(* Logix 5000 project; controller MV vendor 1 type 14 code 217 rev 31.11; software revision 31.00; part 33 of 53 *)
(* tags used below, declared in another part *)
   active : BOOL;
   Alarm_Reset : BOOL;
   CheckTimeMask : INT;
   CLOCK_system_set : BOOL;
   CLOCKsetvalues : DINT[7];
   colon_string : STRING;
   CurrentTime : DateTime;
   CWD : CHECKWORD_FLAGS;
   Default_Check_Time : DINT;
   FtoF_raw_input : REAL;
   FVHR26_3102 : PlantItem;   // Valve FVHR26_31/02
   FVHR26_3102_ALARM : ALARM_DIGITAL;
   FVHR26_3102_CL : ALIAS FOR RIO_Rack_2:14:I.Data.4;   // Valve FVHR26_31/02 Closed
   FVHR26_3102_DR : ALIAS FOR RIO_Rack_2:15:O.Data.18;   // Valve FVHR26_31/02 Drive
   FVHR26_3102_OP : ALIAS FOR RIO_Rack_2:14:I.Data.5;   // Valve FVHR26_31/02 Open
   FVHR26_3103 : PlantItem;   // Valve FVHR26_31/03
   FVHR26_3103_ALARM : ALARM_DIGITAL;
   FVHR26_3103_CL : ALIAS FOR RIO_Rack_2:14:I.Data.6;   // Valve FVHR26_31/03 Closed
   FVHR26_3103_DR : ALIAS FOR RIO_Rack_2:15:O.Data.19;   // Valve FVHR26_31/03 Drive
   FVHR26_3103_OP : ALIAS FOR RIO_Rack_2:14:I.Data.7;   // Valve FVHR26_31/03 Open
   FVHRCH201 : PlantItem;   // Valve FVHRCH201
   FVHRCH201_ALARM : ALARM_DIGITAL;
   FVHRCH201_CL : ALIAS FOR RIO_Rack_2:14:I.Data.10;   // Valve FVHRCH201 Closed
   FVHRCH201_DR : ALIAS FOR RIO_Rack_2:15:O.Data.21;   // Valve FVHRCH201 Drive
   FVHRCH201_OP : ALIAS FOR RIO_Rack_2:14:I.Data.11;   // Valve FVHRCH201 Open
   FVHRCH202 : PlantItem;   // Valve FVHRCH202
   FVHRCH202_ALARM : ALARM_DIGITAL;
   FVHRCH202_CL : ALIAS FOR RIO_Rack_2:14:I.Data.14;   // Valve FVHRCH202 Closed
   FVHRCH202_DR : ALIAS FOR RIO_Rack_2:15:O.Data.23;   // Valve FVHRCH202 Drive
   FVHRCH202_OP : ALIAS FOR RIO_Rack_2:14:I.Data.15;   // Valve FVHRCH202 Open
   FVHRCW01 : PlantItem;   // Valve FVHRCW01
   FVHRCW01_ALARM : ALARM_DIGITAL;
   FVHRCW01_CL : ALIAS FOR RIO_Rack_2:14:I.Data.12;   // Valve FVHRCW01 Closed
   FVHRCW01_DR : ALIAS FOR RIO_Rack_2:15:O.Data.22;   // Valve FVHRCW01 Drive
   FVHRCW01_OP : ALIAS FOR RIO_Rack_2:14:I.Data.13;   // Valve FVHRCW01 Open
   FVHRM01 : PlantItem;   // Valve FVHRM01
   FVHRM01_ALARM : ALARM_DIGITAL;
   FVHRM01_CL : ALIAS FOR RIO_Rack_2:13:I.Data.30;   // Valve FVHRM01 Closed
   FVHRM01_DR : ALIAS FOR RIO_Rack_2:15:O.Data.15;   // Valve FVHRM01 Drive
   FVHRM01_OP : ALIAS FOR RIO_Rack_2:13:I.Data.31;   // Valve FVHRM01 Open
   FVHRM02 : PlantItem;   // Valve FVHRM02
   FVHRM02_ALARM : ALARM_DIGITAL;
   FVHRM02_CL : ALIAS FOR RIO_Rack_2:14:I.Data.0;   // Valve FVHRM02 Closed
   FVHRM02_DR : ALIAS FOR RIO_Rack_2:15:O.Data.16;   // Valve FVHRM02 Drive
   FVHRM02_OP : ALIAS FOR RIO_Rack_2:14:I.Data.1;   // Valve FVHRM02 Open
   FVHRM03 : PlantItem;   // Valve FVHRM03
   FVHRM03_ALARM : ALARM_DIGITAL;
   FVHRM03_CL : ALIAS FOR RIO_Rack_2:14:I.Data.8;   // Valve FVHRM03 Closed
   FVHRM03_DR : ALIAS FOR RIO_Rack_2:15:O.Data.20;   // Valve FVHRM03 Drive
   FVHRM03_OP : ALIAS FOR RIO_Rack_2:14:I.Data.9;   // Valve FVHRM03 Open
   FVHRM04 : PlantItem;   // Valve FVHRM04
   FVHRM04_ALARM : ALARM_DIGITAL;
   FVHRM04_CL : ALIAS FOR RIO_Rack_2:13:I.Data.12;   // Valve FVHRM04 Closed
   FVHRM04_DR : ALIAS FOR RIO_Rack_2:15:O.Data.6;   // Valve FVHRM04 Drive
   FVHRM04_OP : ALIAS FOR RIO_Rack_2:13:I.Data.13;   // Valve FVHRM04 Open
   FVHRMD01 : PlantItem;   // Valve FVHRMD01
   FVHRMD01_ALARM : ALARM_DIGITAL;
   FVHRMD01_CL : ALIAS FOR RIO_Rack_2:13:I.Data.14;   // Valve FVHRMD01 Closed
   FVHRMD01_DR : ALIAS FOR RIO_Rack_2:15:O.Data.7;   // Valve FVHRMD01 Drive
   FVHRMD01_OP : ALIAS FOR RIO_Rack_2:13:I.Data.15;   // Valve FVHRMD01 Open
   hr_string : STRING;
   IGI_TestBit : BOOL;
   Item_Faults_Are_Latched : BOOL;
   Item_Simulation_Flag : BOOL;
   ItoF_raw_input : INT;
   mn_string : STRING;
   MV_DayOfWeek : DINT;
   MV_DayOfWeekONS : BOOL;
   MV_SFile : INT[255];   // SLC Equivalent System File, So Original Code Can Remain
   One_Second_One_Scan : ALIAS FOR One_Second_1_scan;
   result_string : STRING;
   scale_analog_int : DINT;
   scale_analog_result : REAL;
   scale_eu_max : REAL;
   scale_eu_min : REAL;
   scale_raw_input : REAL;
   scale_raw_max : REAL;
   scale_raw_min : REAL;
   scale_routine_active : BOOL;
   scale_temp : REAL;
   se_string : STRING;
   seconds_input_DINT : DINT;
   temp : INT;
   temp_hr : INT;
   temp_mn : INT;
   temp_se : INT;
   zero_string : STRING;
(* MC_Common, continued *)

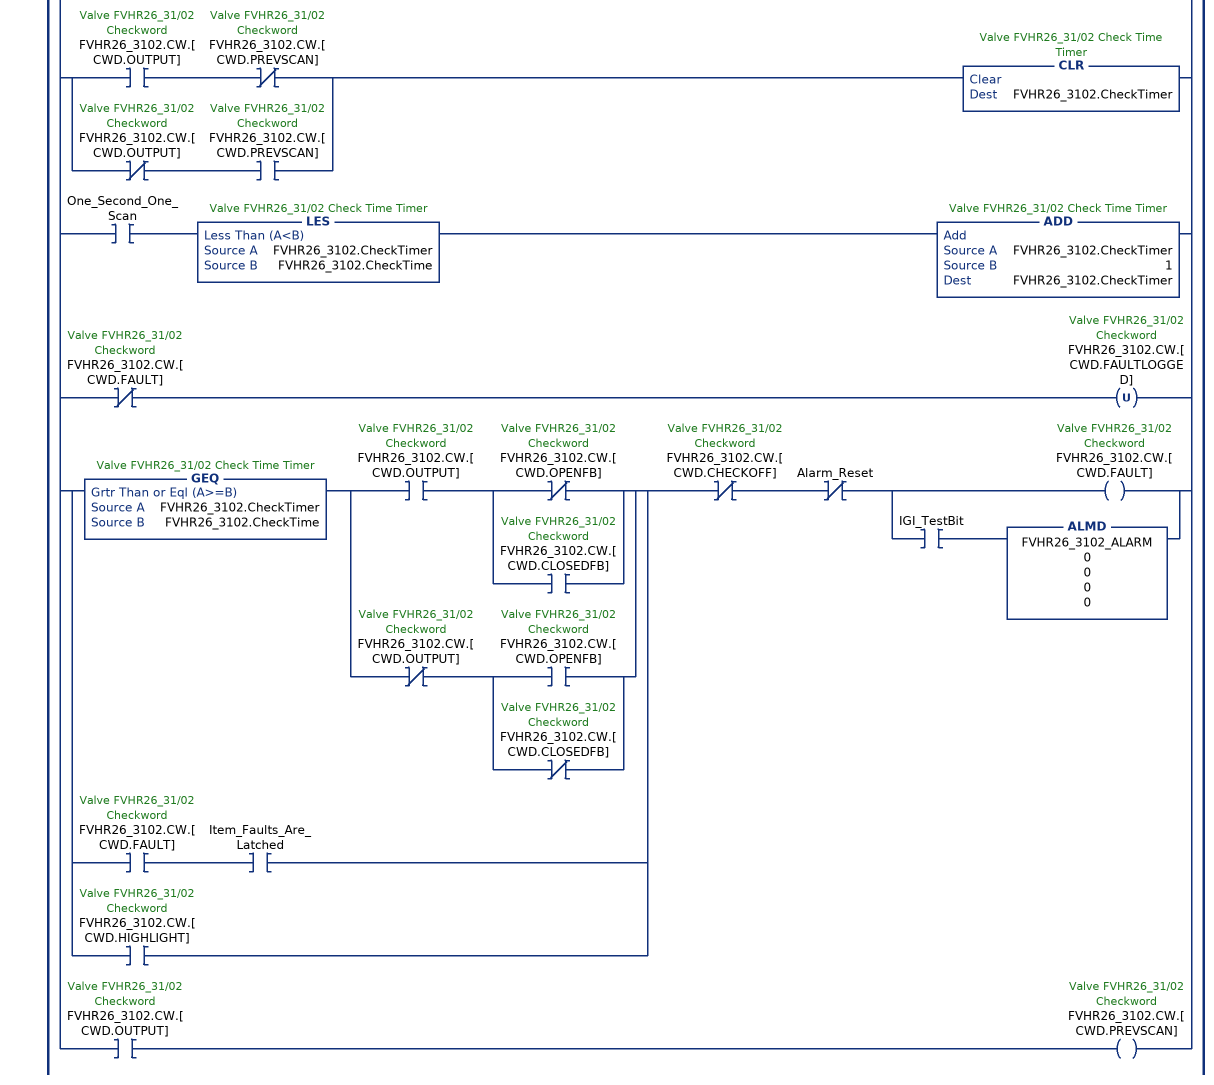
   [picture p757: MC_Common/MC_Valves rungs 79-79]
   79: [NEQ(FVHR26_3102.DriveBits,0) OTE(FVHR26_3102.CW.[CWD.AUTODRV]) ,[XIC(FVHR26_3102.CW.[CWD.AUTODRV]) XIO(FVHR26_3102.CW.[CWD.MANUAL]) ,XIC(FVHR26_3102.CW.[CWD.MANDRV]) XIC(FVHR26_3102.CW.[CWD.MANUAL]) ] OTE(FVHR26_3102.CW.[CWD.OUTPUT]) ,XIC(FVHR26_3102.CW.[CWD.OUTPUT]) OTE(FVHR26_3102_DR) ,XIC(S:FS) [OTU(FVHR26_3102.CW.[CWD.MANUAL]) ,LEQ(FVHR26_3102.CheckTime,0) MOV(Default_Check_Time,FVHR26_3102.CheckTime) ] ,[[XIC(FVHR26_3102_OP) XIO(Item_Simulation_Flag) ,XIC(Item_Simulation_Flag) XIC(FVHR26_3102.CW.[CWD.OUTPUT]) XIO(FVHR26_3102.CW.[CWD.SIMFAIL]) ] OTE(FVHR26_3102.CW.[CWD.OPENFB]) ,[XIC(FVHR26_3102_CL) XIO(Item_Simulation_Flag) ,XIC(Item_Simulation_Flag) XIO(FVHR26_3102.CW.[CWD.OUTPUT]) XIO(FVHR26_3102.CW.[CWD.SIMFAIL]) ] OTE(FVHR26_3102.CW.[CWD.CLOSEDFB]) ] ,[XIC(FVHR26_3102.CW.[CWD.OUTPUT]) XIO(FVHR26_3102.CW.[CWD.PREVSCAN]) ,XIO(FVHR26_3102.CW.[CWD.OUTPUT]) XIC(FVHR26_3102.CW.[CWD.PREVSCAN]) ] CLR(FVHR26_3102.CheckTimer) ,XIC(One_Second_One_Scan) LES(FVHR26_3102.CheckTimer,FVHR26_3102.CheckTime) ADD(FVHR26_3102.CheckTimer,1,FVHR26_3102.CheckTimer) ,XIO(FVHR26_3102.CW.[CWD.FAULT]) OTU(FVHR26_3102.CW.[CWD.FAULTLOGGED]) ,[GEQ(FVHR26_3102.CheckTimer,FVHR26_3102.CheckTime) [XIC(FVHR26_3102.CW.[CWD.OUTPUT]) [XIO(FVHR26_3102.CW.[CWD.OPENFB]) ,XIC(FVHR26_3102.CW.[CWD.CLOSEDFB]) ] ,XIO(FVHR26_3102.CW.[CWD.OUTPUT]) [XIC(FVHR26_3102.CW.[CWD.OPENFB]) ,XIO(FVHR26_3102.CW.[CWD.CLOSEDFB]) ] ] ,XIC(FVHR26_3102.CW.[CWD.FAULT]) XIC(Item_Faults_Are_Latched) ,XIC(FVHR26_3102.CW.[CWD.HIGHLIGHT]) ] XIO(FVHR26_3102.CW.[CWD.CHECKOFF]) XIO(Alarm_Reset) [OTE(FVHR26_3102.CW.[CWD.FAULT]) ,XIC(IGI_TestBit) ALMD(FVHR26_3102_ALARM,0,0,0,0) ] ,XIC(FVHR26_3102.CW.[CWD.OUTPUT]) OTE(FVHR26_3102.CW.[CWD.PREVSCAN]) ];
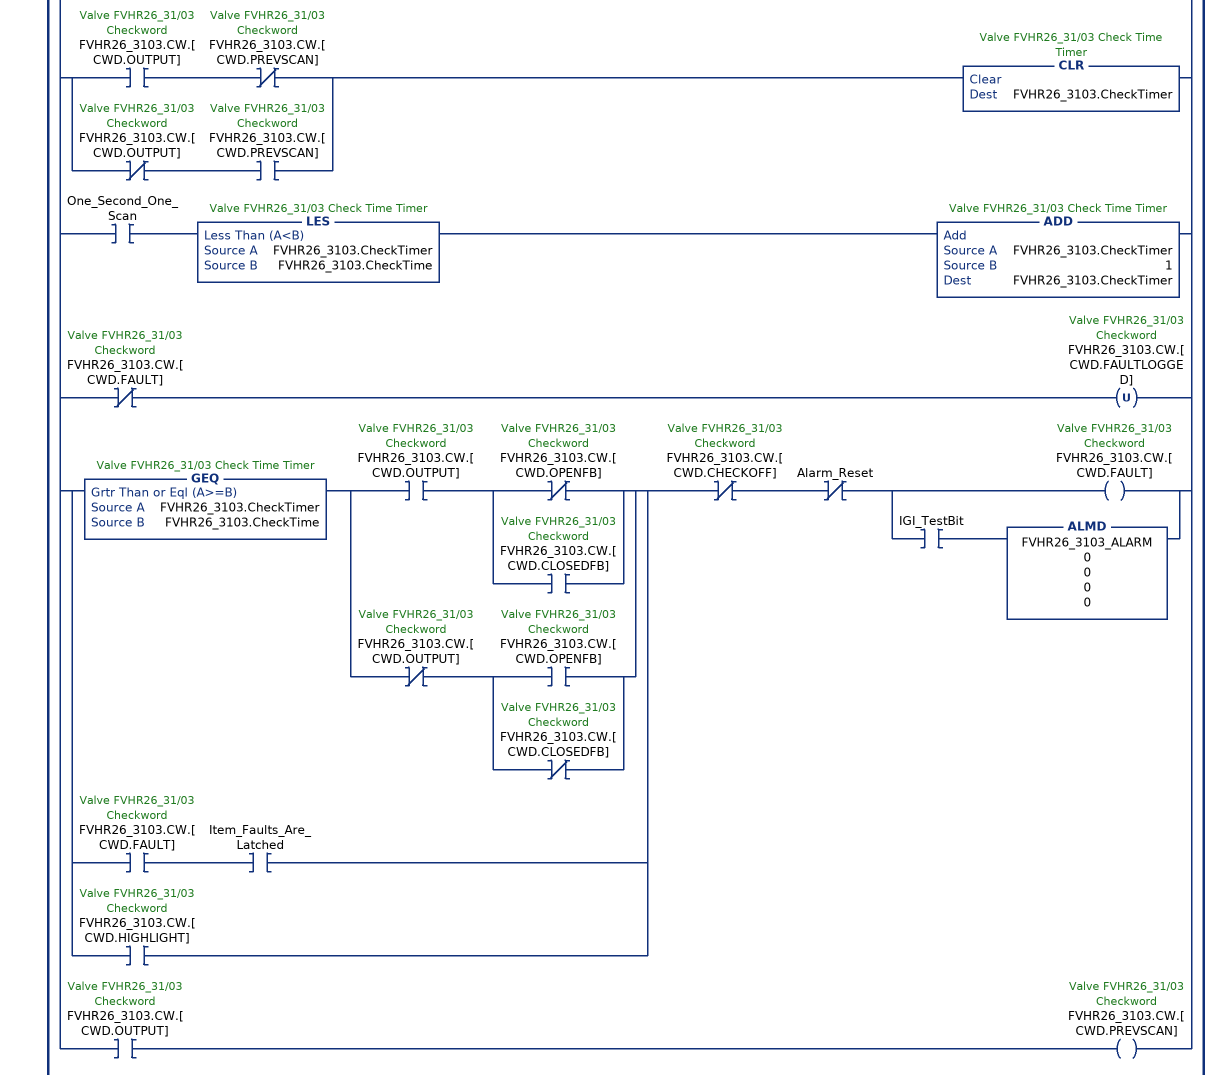
   80: [NEQ(FVHR26_3103.DriveBits,0) OTE(FVHR26_3103.CW.[CWD.AUTODRV]) ,[XIC(FVHR26_3103.CW.[CWD.AUTODRV]) XIO(FVHR26_3103.CW.[CWD.MANUAL]) ,XIC(FVHR26_3103.CW.[CWD.MANDRV]) XIC(FVHR26_3103.CW.[CWD.MANUAL]) ] OTE(FVHR26_3103.CW.[CWD.OUTPUT]) ,XIC(FVHR26_3103.CW.[CWD.OUTPUT]) OTE(FVHR26_3103_DR) ,XIC(S:FS) [OTU(FVHR26_3103.CW.[CWD.MANUAL]) ,LEQ(FVHR26_3103.CheckTime,0) MOV(Default_Check_Time,FVHR26_3103.CheckTime) ] ,[[XIC(FVHR26_3103_OP) XIO(Item_Simulation_Flag) ,XIC(Item_Simulation_Flag) XIC(FVHR26_3103.CW.[CWD.OUTPUT]) XIO(FVHR26_3103.CW.[CWD.SIMFAIL]) ] OTE(FVHR26_3103.CW.[CWD.OPENFB]) ,[XIC(FVHR26_3103_CL) XIO(Item_Simulation_Flag) ,XIC(Item_Simulation_Flag) XIO(FVHR26_3103.CW.[CWD.OUTPUT]) XIO(FVHR26_3103.CW.[CWD.SIMFAIL]) ] OTE(FVHR26_3103.CW.[CWD.CLOSEDFB]) ] ,[XIC(FVHR26_3103.CW.[CWD.OUTPUT]) XIO(FVHR26_3103.CW.[CWD.PREVSCAN]) ,XIO(FVHR26_3103.CW.[CWD.OUTPUT]) XIC(FVHR26_3103.CW.[CWD.PREVSCAN]) ] CLR(FVHR26_3103.CheckTimer) ,XIC(One_Second_One_Scan) LES(FVHR26_3103.CheckTimer,FVHR26_3103.CheckTime) ADD(FVHR26_3103.CheckTimer,1,FVHR26_3103.CheckTimer) ,XIO(FVHR26_3103.CW.[CWD.FAULT]) OTU(FVHR26_3103.CW.[CWD.FAULTLOGGED]) ,[GEQ(FVHR26_3103.CheckTimer,FVHR26_3103.CheckTime) [XIC(FVHR26_3103.CW.[CWD.OUTPUT]) [XIO(FVHR26_3103.CW.[CWD.OPENFB]) ,XIC(FVHR26_3103.CW.[CWD.CLOSEDFB]) ] ,XIO(FVHR26_3103.CW.[CWD.OUTPUT]) [XIC(FVHR26_3103.CW.[CWD.OPENFB]) ,XIO(FVHR26_3103.CW.[CWD.CLOSEDFB]) ] ] ,XIC(FVHR26_3103.CW.[CWD.FAULT]) XIC(Item_Faults_Are_Latched) ,XIC(FVHR26_3103.CW.[CWD.HIGHLIGHT]) ] XIO(FVHR26_3103.CW.[CWD.CHECKOFF]) XIO(Alarm_Reset) [OTE(FVHR26_3103.CW.[CWD.FAULT]) ,XIC(IGI_TestBit) ALMD(FVHR26_3103_ALARM,0,0,0,0) ] ,XIC(FVHR26_3103.CW.[CWD.OUTPUT]) OTE(FVHR26_3103.CW.[CWD.PREVSCAN]) ];
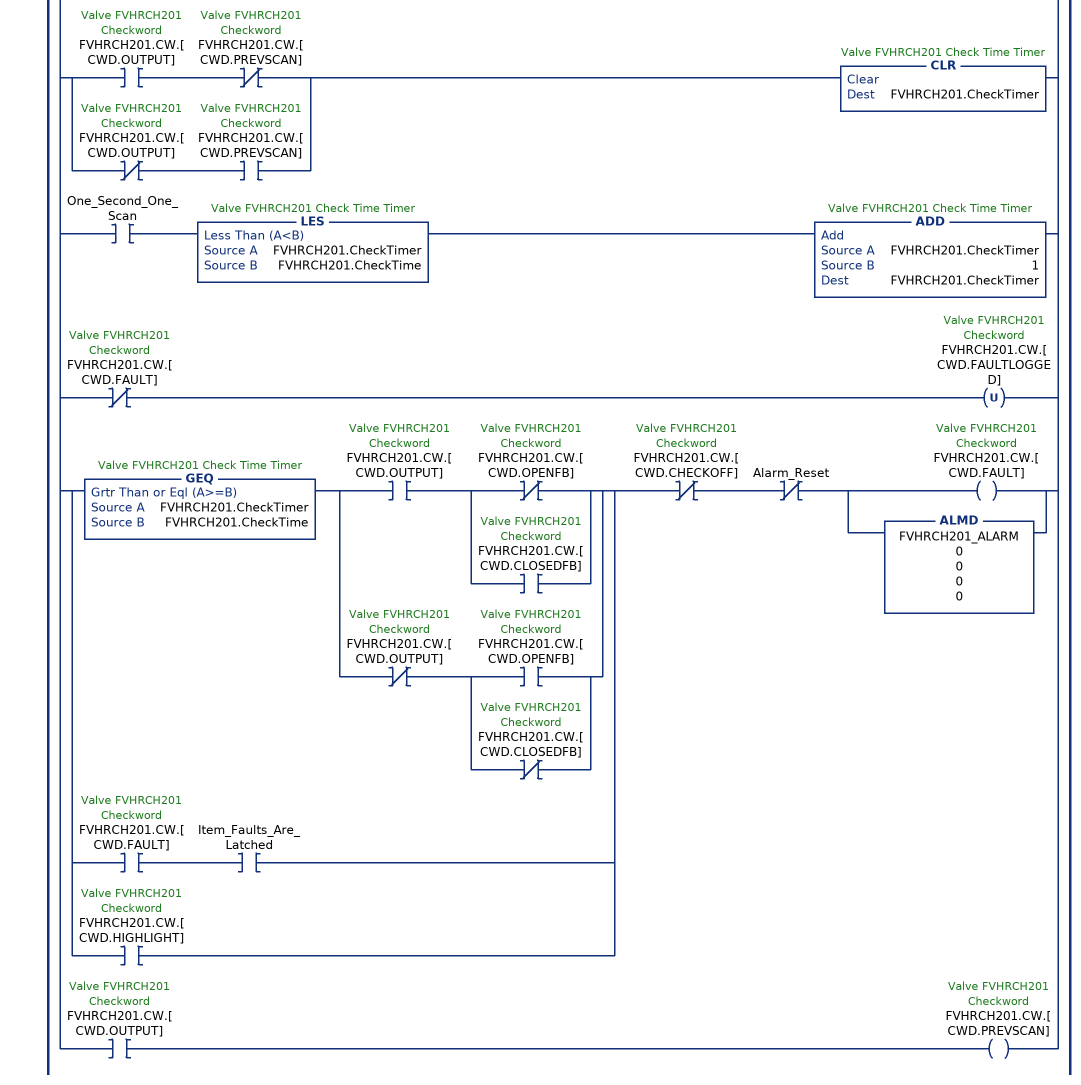
   81: [NEQ(FVHRCH201.DriveBits,0) OTE(FVHRCH201.CW.[CWD.AUTODRV]) ,[XIC(FVHRCH201.CW.[CWD.AUTODRV]) XIO(FVHRCH201.CW.[CWD.MANUAL]) ,XIC(FVHRCH201.CW.[CWD.MANDRV]) XIC(FVHRCH201.CW.[CWD.MANUAL]) ] OTE(FVHRCH201.CW.[CWD.OUTPUT]) ,XIC(FVHRCH201.CW.[CWD.OUTPUT]) OTE(FVHRCH201_DR) ,XIC(S:FS) [OTU(FVHRCH201.CW.[CWD.MANUAL]) ,LEQ(FVHRCH201.CheckTime,0) MOV(Default_Check_Time,FVHRCH201.CheckTime) ] ,[[XIC(FVHRCH201_OP) XIO(Item_Simulation_Flag) ,XIC(Item_Simulation_Flag) XIC(FVHRCH201.CW.[CWD.OUTPUT]) XIO(FVHRCH201.CW.[CWD.SIMFAIL]) ] OTE(FVHRCH201.CW.[CWD.OPENFB]) ,[XIC(FVHRCH201_CL) XIO(Item_Simulation_Flag) ,XIC(Item_Simulation_Flag) XIO(FVHRCH201.CW.[CWD.OUTPUT]) XIO(FVHRCH201.CW.[CWD.SIMFAIL]) ] OTE(FVHRCH201.CW.[CWD.CLOSEDFB]) ] ,[XIC(FVHRCH201.CW.[CWD.OUTPUT]) XIO(FVHRCH201.CW.[CWD.PREVSCAN]) ,XIO(FVHRCH201.CW.[CWD.OUTPUT]) XIC(FVHRCH201.CW.[CWD.PREVSCAN]) ] CLR(FVHRCH201.CheckTimer) ,XIC(One_Second_One_Scan) LES(FVHRCH201.CheckTimer,FVHRCH201.CheckTime) ADD(FVHRCH201.CheckTimer,1,FVHRCH201.CheckTimer) ,XIO(FVHRCH201.CW.[CWD.FAULT]) OTU(FVHRCH201.CW.[CWD.FAULTLOGGED]) ,[GEQ(FVHRCH201.CheckTimer,FVHRCH201.CheckTime) [XIC(FVHRCH201.CW.[CWD.OUTPUT]) [XIO(FVHRCH201.CW.[CWD.OPENFB]) ,XIC(FVHRCH201.CW.[CWD.CLOSEDFB]) ] ,XIO(FVHRCH201.CW.[CWD.OUTPUT]) [XIC(FVHRCH201.CW.[CWD.OPENFB]) ,XIO(FVHRCH201.CW.[CWD.CLOSEDFB]) ] ] ,XIC(FVHRCH201.CW.[CWD.FAULT]) XIC(Item_Faults_Are_Latched) ,XIC(FVHRCH201.CW.[CWD.HIGHLIGHT]) ] XIO(FVHRCH201.CW.[CWD.CHECKOFF]) XIO(Alarm_Reset) [OTE(FVHRCH201.CW.[CWD.FAULT]) ,ALMD(FVHRCH201_ALARM,0,0,0,0) ] ,XIC(FVHRCH201.CW.[CWD.OUTPUT]) OTE(FVHRCH201.CW.[CWD.PREVSCAN]) ];
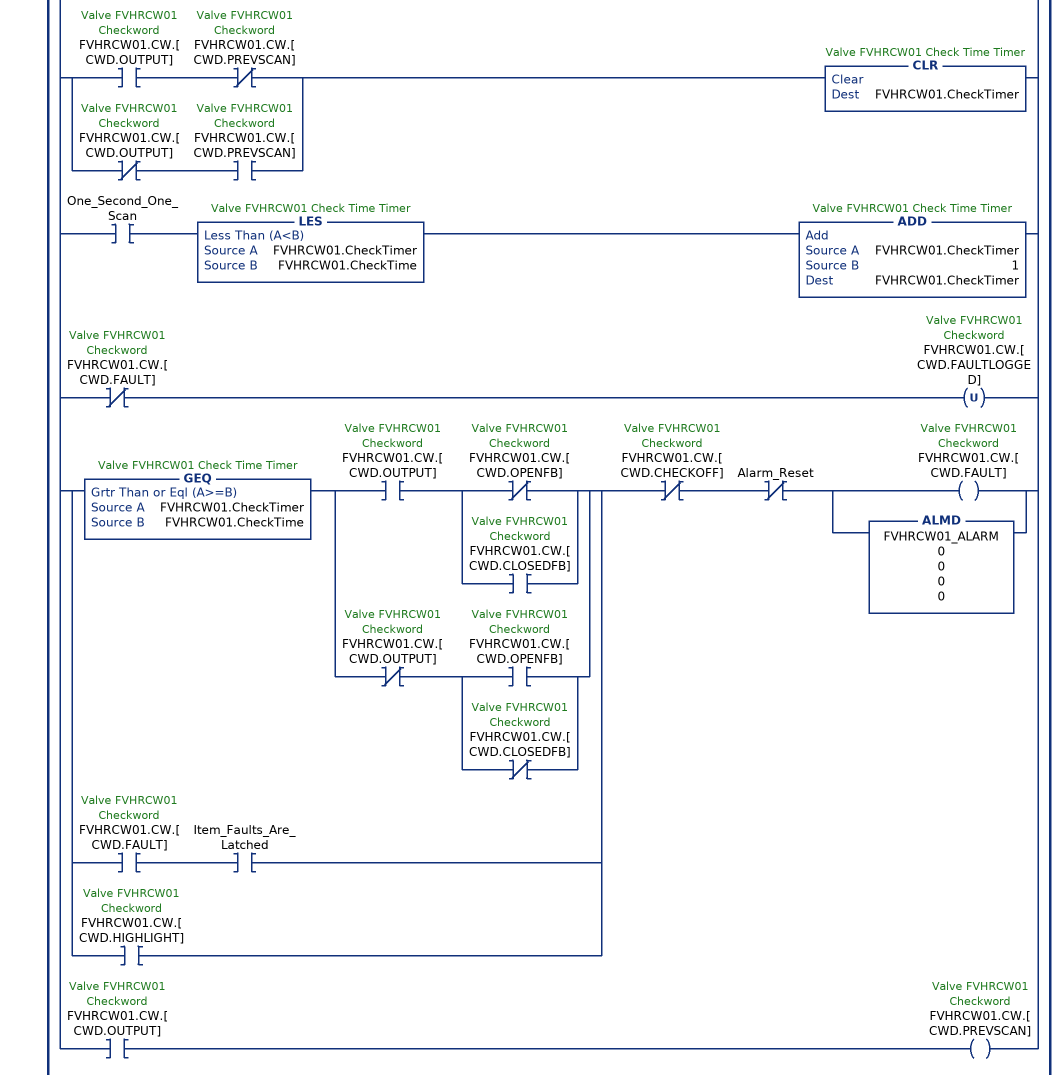
   82: [NEQ(FVHRCW01.DriveBits,0) OTE(FVHRCW01.CW.[CWD.AUTODRV]) ,[XIC(FVHRCW01.CW.[CWD.AUTODRV]) XIO(FVHRCW01.CW.[CWD.MANUAL]) ,XIC(FVHRCW01.CW.[CWD.MANDRV]) XIC(FVHRCW01.CW.[CWD.MANUAL]) ] OTE(FVHRCW01.CW.[CWD.OUTPUT]) ,XIC(FVHRCW01.CW.[CWD.OUTPUT]) OTE(FVHRCW01_DR) ,XIC(S:FS) [OTU(FVHRCW01.CW.[CWD.MANUAL]) ,LEQ(FVHRCW01.CheckTime,0) MOV(Default_Check_Time,FVHRCW01.CheckTime) ] ,[[XIC(FVHRCW01_OP) XIO(Item_Simulation_Flag) ,XIC(Item_Simulation_Flag) XIC(FVHRCW01.CW.[CWD.OUTPUT]) XIO(FVHRCW01.CW.[CWD.SIMFAIL]) ] OTE(FVHRCW01.CW.[CWD.OPENFB]) ,[XIC(FVHRCW01_CL) XIO(Item_Simulation_Flag) ,XIC(Item_Simulation_Flag) XIO(FVHRCW01.CW.[CWD.OUTPUT]) XIO(FVHRCW01.CW.[CWD.SIMFAIL]) ] OTE(FVHRCW01.CW.[CWD.CLOSEDFB]) ] ,[XIC(FVHRCW01.CW.[CWD.OUTPUT]) XIO(FVHRCW01.CW.[CWD.PREVSCAN]) ,XIO(FVHRCW01.CW.[CWD.OUTPUT]) XIC(FVHRCW01.CW.[CWD.PREVSCAN]) ] CLR(FVHRCW01.CheckTimer) ,XIC(One_Second_One_Scan) LES(FVHRCW01.CheckTimer,FVHRCW01.CheckTime) ADD(FVHRCW01.CheckTimer,1,FVHRCW01.CheckTimer) ,XIO(FVHRCW01.CW.[CWD.FAULT]) OTU(FVHRCW01.CW.[CWD.FAULTLOGGED]) ,[GEQ(FVHRCW01.CheckTimer,FVHRCW01.CheckTime) [XIC(FVHRCW01.CW.[CWD.OUTPUT]) [XIO(FVHRCW01.CW.[CWD.OPENFB]) ,XIC(FVHRCW01.CW.[CWD.CLOSEDFB]) ] ,XIO(FVHRCW01.CW.[CWD.OUTPUT]) [XIC(FVHRCW01.CW.[CWD.OPENFB]) ,XIO(FVHRCW01.CW.[CWD.CLOSEDFB]) ] ] ,XIC(FVHRCW01.CW.[CWD.FAULT]) XIC(Item_Faults_Are_Latched) ,XIC(FVHRCW01.CW.[CWD.HIGHLIGHT]) ] XIO(FVHRCW01.CW.[CWD.CHECKOFF]) XIO(Alarm_Reset) [OTE(FVHRCW01.CW.[CWD.FAULT]) ,ALMD(FVHRCW01_ALARM,0,0,0,0) ] ,XIC(FVHRCW01.CW.[CWD.OUTPUT]) OTE(FVHRCW01.CW.[CWD.PREVSCAN]) ];
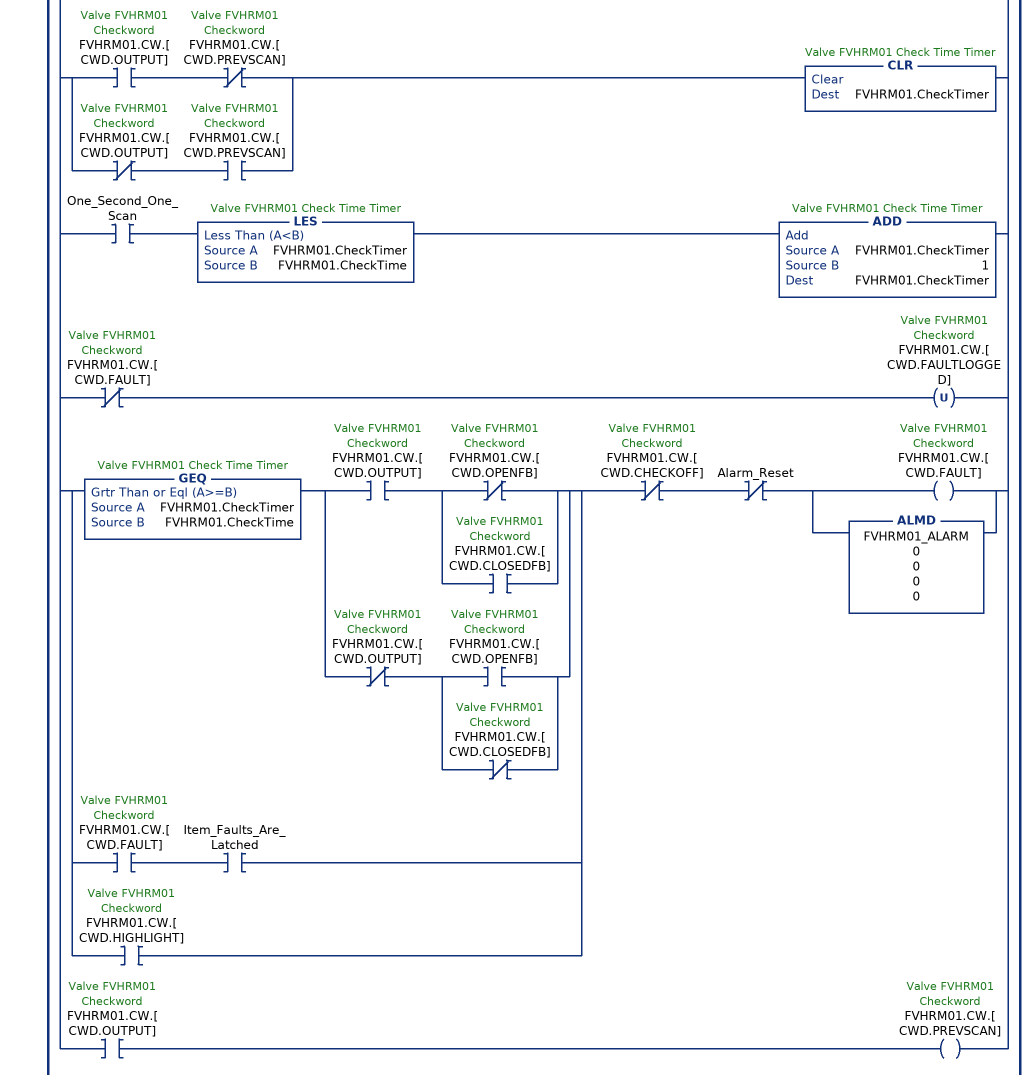
   83: [NEQ(FVHRM01.DriveBits,0) OTE(FVHRM01.CW.[CWD.AUTODRV]) ,[XIC(FVHRM01.CW.[CWD.AUTODRV]) XIO(FVHRM01.CW.[CWD.MANUAL]) ,XIC(FVHRM01.CW.[CWD.MANDRV]) XIC(FVHRM01.CW.[CWD.MANUAL]) ] OTE(FVHRM01.CW.[CWD.OUTPUT]) ,XIC(FVHRM01.CW.[CWD.OUTPUT]) OTE(FVHRM01_DR) ,XIC(S:FS) [OTU(FVHRM01.CW.[CWD.MANUAL]) ,LEQ(FVHRM01.CheckTime,0) MOV(Default_Check_Time,FVHRM01.CheckTime) ] ,[[XIC(FVHRM01_OP) XIO(Item_Simulation_Flag) ,XIC(Item_Simulation_Flag) XIC(FVHRM01.CW.[CWD.OUTPUT]) XIO(FVHRM01.CW.[CWD.SIMFAIL]) ] OTE(FVHRM01.CW.[CWD.OPENFB]) ,[XIC(FVHRM01_CL) XIO(Item_Simulation_Flag) ,XIC(Item_Simulation_Flag) XIO(FVHRM01.CW.[CWD.OUTPUT]) XIO(FVHRM01.CW.[CWD.SIMFAIL]) ] OTE(FVHRM01.CW.[CWD.CLOSEDFB]) ] ,[XIC(FVHRM01.CW.[CWD.OUTPUT]) XIO(FVHRM01.CW.[CWD.PREVSCAN]) ,XIO(FVHRM01.CW.[CWD.OUTPUT]) XIC(FVHRM01.CW.[CWD.PREVSCAN]) ] CLR(FVHRM01.CheckTimer) ,XIC(One_Second_One_Scan) LES(FVHRM01.CheckTimer,FVHRM01.CheckTime) ADD(FVHRM01.CheckTimer,1,FVHRM01.CheckTimer) ,XIO(FVHRM01.CW.[CWD.FAULT]) OTU(FVHRM01.CW.[CWD.FAULTLOGGED]) ,[GEQ(FVHRM01.CheckTimer,FVHRM01.CheckTime) [XIC(FVHRM01.CW.[CWD.OUTPUT]) [XIO(FVHRM01.CW.[CWD.OPENFB]) ,XIC(FVHRM01.CW.[CWD.CLOSEDFB]) ] ,XIO(FVHRM01.CW.[CWD.OUTPUT]) [XIC(FVHRM01.CW.[CWD.OPENFB]) ,XIO(FVHRM01.CW.[CWD.CLOSEDFB]) ] ] ,XIC(FVHRM01.CW.[CWD.FAULT]) XIC(Item_Faults_Are_Latched) ,XIC(FVHRM01.CW.[CWD.HIGHLIGHT]) ] XIO(FVHRM01.CW.[CWD.CHECKOFF]) XIO(Alarm_Reset) [OTE(FVHRM01.CW.[CWD.FAULT]) ,ALMD(FVHRM01_ALARM,0,0,0,0) ] ,XIC(FVHRM01.CW.[CWD.OUTPUT]) OTE(FVHRM01.CW.[CWD.PREVSCAN]) ];
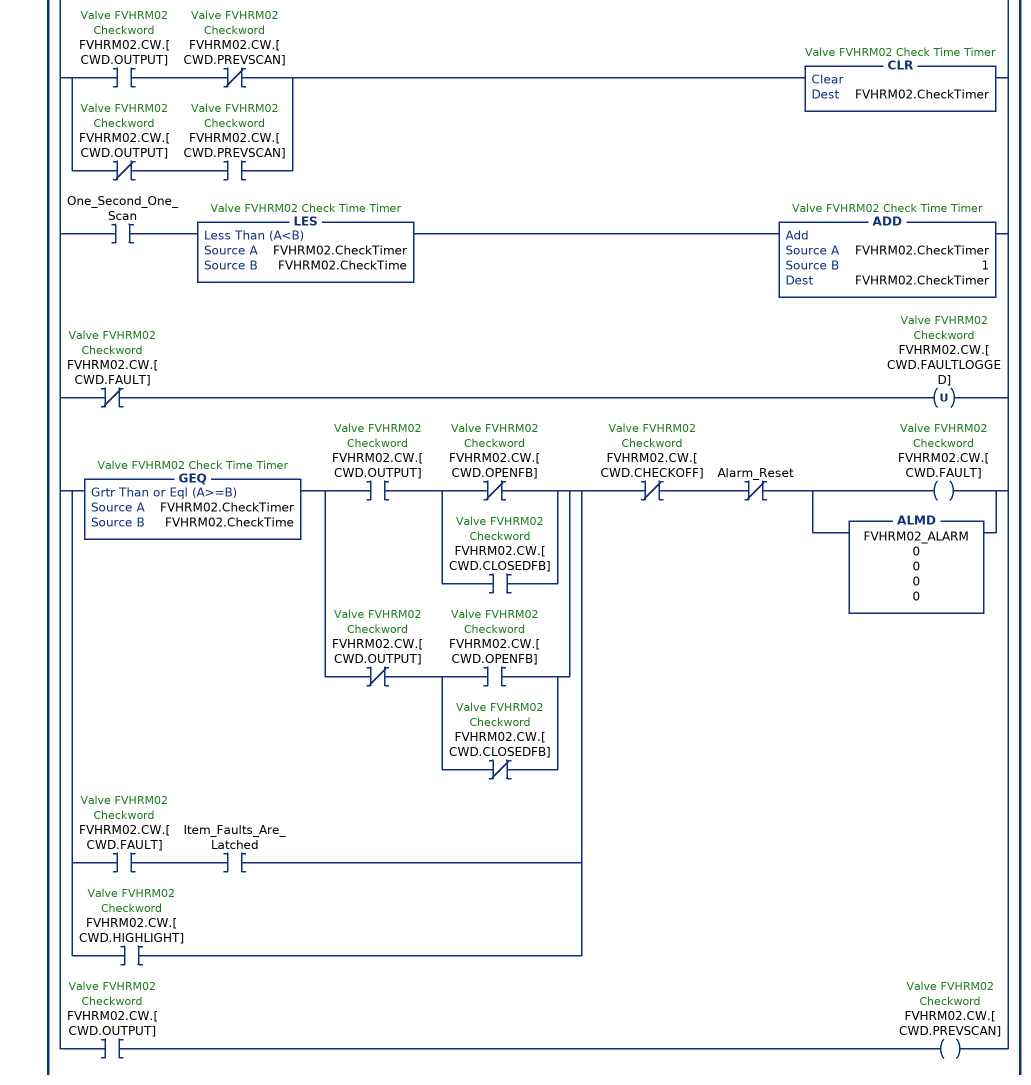
   84: [NEQ(FVHRM02.DriveBits,0) OTE(FVHRM02.CW.[CWD.AUTODRV]) ,[XIC(FVHRM02.CW.[CWD.AUTODRV]) XIO(FVHRM02.CW.[CWD.MANUAL]) ,XIC(FVHRM02.CW.[CWD.MANDRV]) XIC(FVHRM02.CW.[CWD.MANUAL]) ] OTE(FVHRM02.CW.[CWD.OUTPUT]) ,XIC(FVHRM02.CW.[CWD.OUTPUT]) OTE(FVHRM02_DR) ,XIC(S:FS) [OTU(FVHRM02.CW.[CWD.MANUAL]) ,LEQ(FVHRM02.CheckTime,0) MOV(Default_Check_Time,FVHRM02.CheckTime) ] ,[[XIC(FVHRM02_OP) XIO(Item_Simulation_Flag) ,XIC(Item_Simulation_Flag) XIC(FVHRM02.CW.[CWD.OUTPUT]) XIO(FVHRM02.CW.[CWD.SIMFAIL]) ] OTE(FVHRM02.CW.[CWD.OPENFB]) ,[XIC(FVHRM02_CL) XIO(Item_Simulation_Flag) ,XIC(Item_Simulation_Flag) XIO(FVHRM02.CW.[CWD.OUTPUT]) XIO(FVHRM02.CW.[CWD.SIMFAIL]) ] OTE(FVHRM02.CW.[CWD.CLOSEDFB]) ] ,[XIC(FVHRM02.CW.[CWD.OUTPUT]) XIO(FVHRM02.CW.[CWD.PREVSCAN]) ,XIO(FVHRM02.CW.[CWD.OUTPUT]) XIC(FVHRM02.CW.[CWD.PREVSCAN]) ] CLR(FVHRM02.CheckTimer) ,XIC(One_Second_One_Scan) LES(FVHRM02.CheckTimer,FVHRM02.CheckTime) ADD(FVHRM02.CheckTimer,1,FVHRM02.CheckTimer) ,XIO(FVHRM02.CW.[CWD.FAULT]) OTU(FVHRM02.CW.[CWD.FAULTLOGGED]) ,[GEQ(FVHRM02.CheckTimer,FVHRM02.CheckTime) [XIC(FVHRM02.CW.[CWD.OUTPUT]) [XIO(FVHRM02.CW.[CWD.OPENFB]) ,XIC(FVHRM02.CW.[CWD.CLOSEDFB]) ] ,XIO(FVHRM02.CW.[CWD.OUTPUT]) [XIC(FVHRM02.CW.[CWD.OPENFB]) ,XIO(FVHRM02.CW.[CWD.CLOSEDFB]) ] ] ,XIC(FVHRM02.CW.[CWD.FAULT]) XIC(Item_Faults_Are_Latched) ,XIC(FVHRM02.CW.[CWD.HIGHLIGHT]) ] XIO(FVHRM02.CW.[CWD.CHECKOFF]) XIO(Alarm_Reset) [OTE(FVHRM02.CW.[CWD.FAULT]) ,ALMD(FVHRM02_ALARM,0,0,0,0) ] ,XIC(FVHRM02.CW.[CWD.OUTPUT]) OTE(FVHRM02.CW.[CWD.PREVSCAN]) ];